VERSION : 0.1
   VAR_INPUT
      Zone : Int;
      ZonePos : Int;
      ClearOfStopDist : Int;
   END_VAR
   VAR_OUTPUT
      CarrierNumber : Int;
      MoveFwdCommand : Bool;
      DriveCmdSpeed : Int;
      NextCarrierNum : Word;
      NextStopPosition : DWord;
      AtCmdPosition : Bool;
      CarrierInTransitToNextZone : Bool;
   END_VAR
   VAR
      PreviousCarrierNumMemory : Word;
      TrafficCopCarrierZnBuffer : Array[0..40] of "UDT_TrafficCop";
      LastCarrierNextZnPos : Int;
      CarNumZnPos : Int;
      NextZone : Int;
      EndPos_LowLimit : DWord;
      EndPos_HighLimit : DWord;
      ClrOfStopPos_LowLimit : DWord;
      ClrOfStopPos_HighLimit : DWord;
      ClearOfStopPos : DWord;
      ClearToMoveTrain : Bool;
      PrevZone : Int;
      PrevZone_CarrierReady : Bool;
      LastCarrierCurrentZnPos : Int;
      LastCarrierNumber : Word;
      CarrierInTransitToProdZone : Bool;
      ResetCarrierInTransToProd : Bool;
      WaitPositionMemory : DInt;
      OneShot : Bool;
      NextCarrierOffset : DWord;
      PrevZone_EndPos_LowLimit : DWord;
      PrevZone_EndPos_HighLimit : DWord;
   END_VAR
   VAR_TEMP
      NextZoneBuffer : Int;
      LastZone : Int;
      HighSpeedSetpoint : Word;
      LowSpeedSetpoint : Word;
      NextZonePosition : Int;
      NextCarrierOffsetSetup1 : UDInt;
      NextCarrierOffsetSetup2 : UDInt;
   END_VAR
   VAR_TEMP   // added for the SCL form of the ladder/FBD networks
      _w1 : Bool;
      _w2 : Bool;
      _w3 : Bool;
      _w4 : Bool;
      _w5 : Bool;
   END_VAR
BEGIN

REGION Network 1
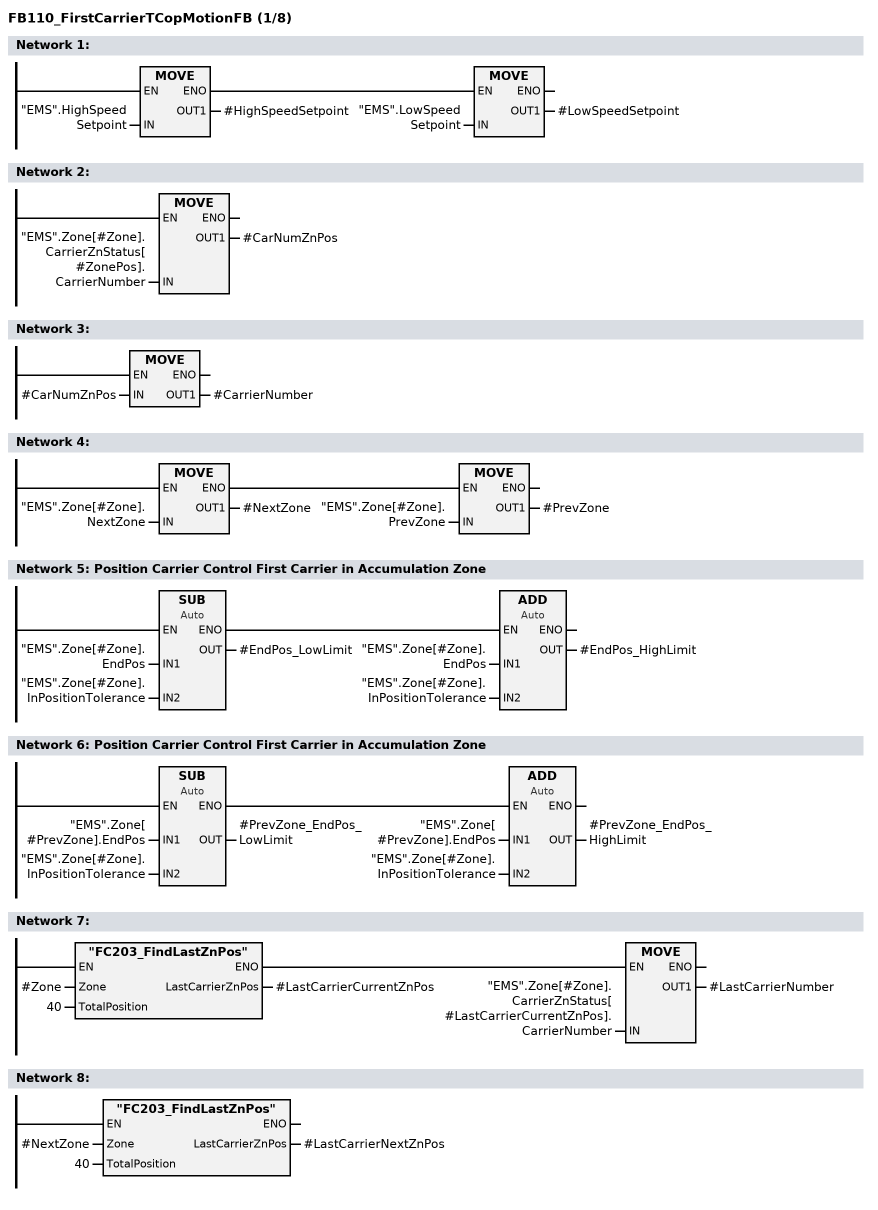
   RUNG wire#powerrail
      Move(in := "EMS".HighSpeedSetpoint, out1 => #HighSpeedSetpoint)
      Move(in := "EMS".LowSpeedSetpoint, out1 => #LowSpeedSetpoint)
   END_RUNG
   // the same network as SCL:
   #HighSpeedSetpoint := "EMS".HighSpeedSetpoint;
   #LowSpeedSetpoint := "EMS".LowSpeedSetpoint;
END_REGION

REGION Network 2
   RUNG wire#powerrail
      Move(in := "EMS".Zone[#Zone].CarrierZnStatus[#ZonePos].CarrierNumber, out1 => #CarNumZnPos)
   END_RUNG
   // the same network as SCL:
   #CarNumZnPos := "EMS".Zone[#Zone].CarrierZnStatus[#ZonePos].CarrierNumber;
END_REGION

REGION Network 3
   RUNG wire#powerrail
      Move(in := #CarNumZnPos, out1 => #CarrierNumber)
   END_RUNG
   // the same network as SCL:
   #CarrierNumber := #CarNumZnPos;
END_REGION

REGION Network 4
   RUNG wire#powerrail
      Move(in := "EMS".Zone[#Zone].NextZone, out1 => #NextZone)
      Move(in := "EMS".Zone[#Zone].PrevZone, out1 => #PrevZone)
   END_RUNG
   // the same network as SCL:
   #NextZone := "EMS".Zone[#Zone].NextZone;
   #PrevZone := "EMS".Zone[#Zone].PrevZone;
END_REGION

REGION Network 5: Position Carrier Control First Carrier in Accumulation Zone
   RUNG wire#powerrail
      Sub(in1 := "EMS".Zone[#Zone].EndPos, in2 := "EMS".Zone[#Zone].InPositionTolerance, out => #EndPos_LowLimit)
      Add(in1 := "EMS".Zone[#Zone].EndPos, in2 := "EMS".Zone[#Zone].InPositionTolerance, out => #EndPos_HighLimit)
   END_RUNG
   // the same network as SCL:
   #EndPos_LowLimit := "EMS".Zone[#Zone].EndPos - "EMS".Zone[#Zone].InPositionTolerance;
   #EndPos_HighLimit := "EMS".Zone[#Zone].EndPos + "EMS".Zone[#Zone].InPositionTolerance;
END_REGION

REGION Network 6: Position Carrier Control First Carrier in Accumulation Zone
   RUNG wire#powerrail
      Sub(in1 := "EMS".Zone[#PrevZone].EndPos, in2 := "EMS".Zone[#Zone].InPositionTolerance, out => #PrevZone_EndPos_LowLimit)
      Add(in1 := "EMS".Zone[#PrevZone].EndPos, in2 := "EMS".Zone[#Zone].InPositionTolerance, out => #PrevZone_EndPos_HighLimit)
   END_RUNG
   // the same network as SCL:
   #PrevZone_EndPos_LowLimit := "EMS".Zone[#PrevZone].EndPos - "EMS".Zone[#Zone].InPositionTolerance;
   #PrevZone_EndPos_HighLimit := "EMS".Zone[#PrevZone].EndPos + "EMS".Zone[#Zone].InPositionTolerance;
END_REGION

REGION Network 7
   RUNG wire#powerrail
      "FC203_FindLastZnPos"(Zone := #Zone, TotalPosition := 40, LastCarrierZnPos => #LastCarrierCurrentZnPos)
      Move(in := "EMS".Zone[#Zone].CarrierZnStatus[#LastCarrierCurrentZnPos].CarrierNumber, out1 => #LastCarrierNumber)
   END_RUNG
   // the same network as SCL:
   "FC203_FindLastZnPos"(Zone := #Zone,
                         TotalPosition := 40,
                         LastCarrierZnPos => #LastCarrierCurrentZnPos,
                         ENO => #_w1);
   IF #_w1 THEN
       #LastCarrierNumber := "EMS".Zone[#Zone].CarrierZnStatus[#LastCarrierCurrentZnPos].CarrierNumber;
   END_IF;
END_REGION

REGION Network 8
   RUNG wire#powerrail
      "FC203_FindLastZnPos"(Zone := #NextZone, TotalPosition := 40, LastCarrierZnPos => #LastCarrierNextZnPos)
   END_RUNG
   // the same network as SCL:
   "FC203_FindLastZnPos"(Zone := #NextZone, TotalPosition := 40, LastCarrierZnPos => #LastCarrierNextZnPos);
END_REGION

REGION Network 9: Position Carrier Control First Carrier in Production Zone
   // Control of First Carrier in Zone Closest to end position/Stop.  Move command is issued to carrier. Carrier will move in auto.
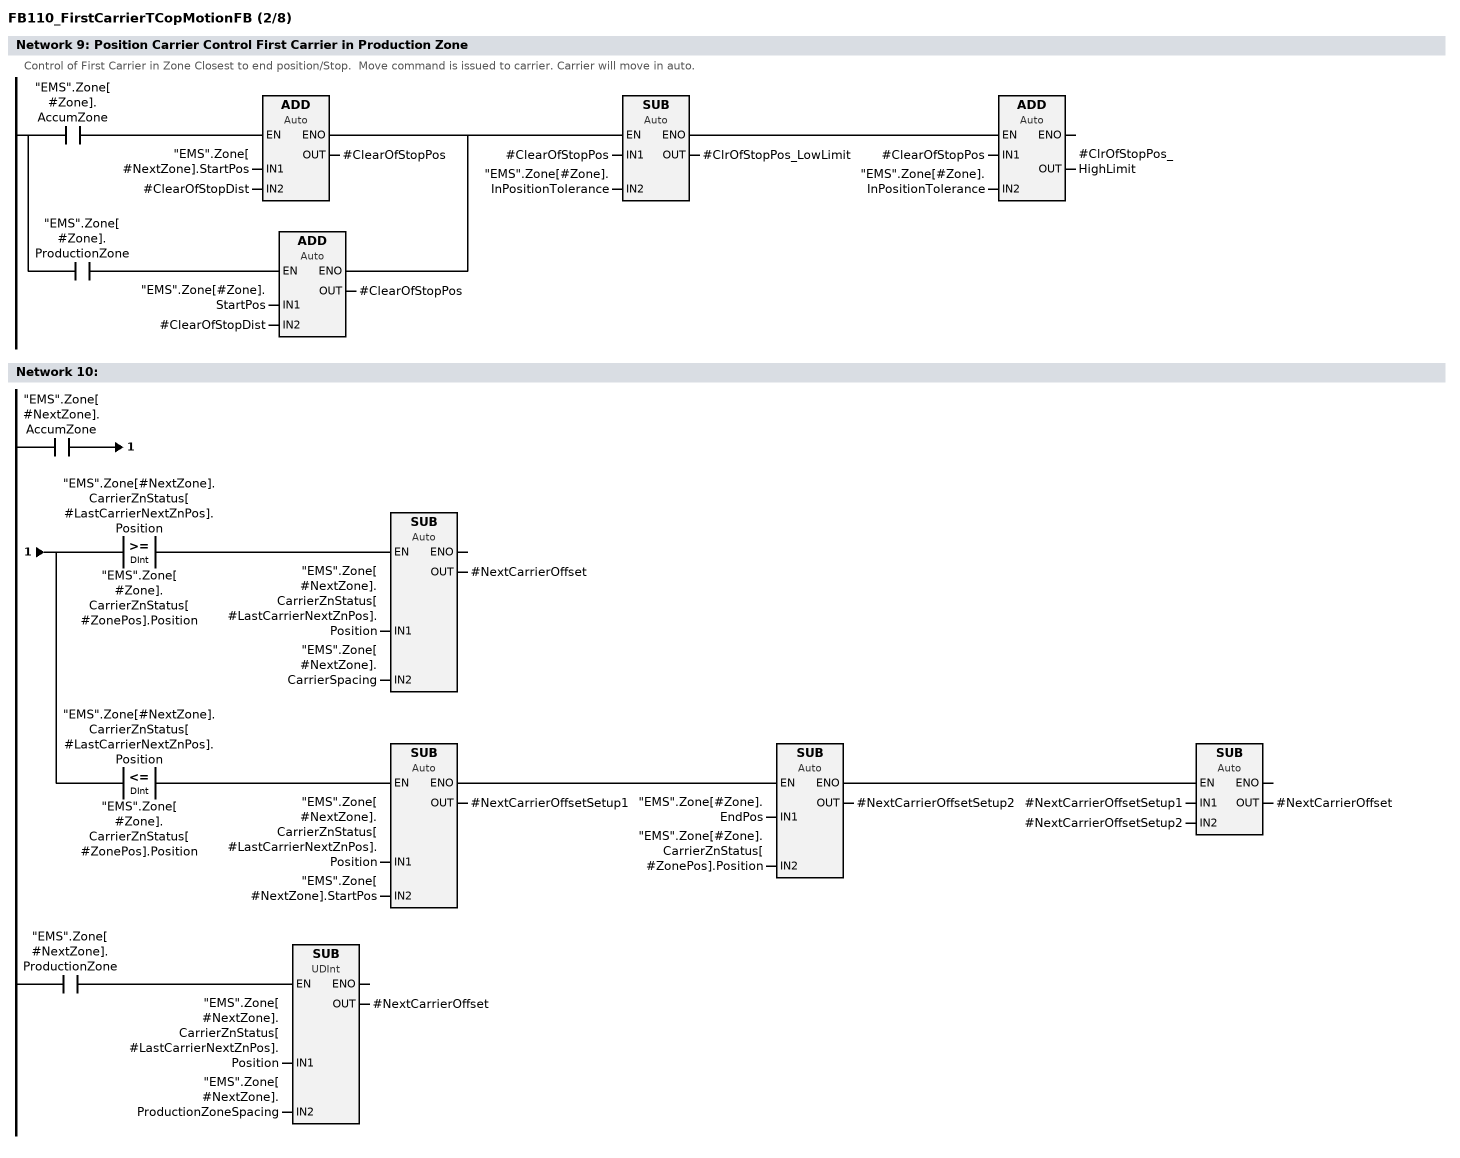
   RUNG wire#powerrail
      Contact( "EMS".Zone[#Zone].AccumZone )
      Add(in1 := "EMS".Zone[#NextZone].StartPos, in2 := #ClearOfStopDist, out => #ClearOfStopPos)
      wire#w1
      Sub(in1 := #ClearOfStopPos, in2 := "EMS".Zone[#Zone].InPositionTolerance, out => #ClrOfStopPos_LowLimit)
      Add(in1 := #ClearOfStopPos, in2 := "EMS".Zone[#Zone].InPositionTolerance, out => #ClrOfStopPos_HighLimit)
   END_RUNG
   RUNG wire#powerrail
      Contact( "EMS".Zone[#Zone].ProductionZone )
      Add(in1 := "EMS".Zone[#Zone].StartPos, in2 := #ClearOfStopDist, out => #ClearOfStopPos)
   END_RUNG wire#w1
   // the same network as SCL:
   IF "EMS".Zone[#Zone].AccumZone THEN
       #ClearOfStopPos := "EMS".Zone[#NextZone].StartPos + #ClearOfStopDist;
   END_IF;
   IF "EMS".Zone[#Zone].ProductionZone THEN
       #ClearOfStopPos := "EMS".Zone[#Zone].StartPos + #ClearOfStopDist;
   END_IF;
   IF "EMS".Zone[#Zone].AccumZone OR "EMS".Zone[#Zone].ProductionZone THEN
       #ClrOfStopPos_LowLimit := #ClearOfStopPos - "EMS".Zone[#Zone].InPositionTolerance;
       #ClrOfStopPos_HighLimit := #ClearOfStopPos + "EMS".Zone[#Zone].InPositionTolerance;
   END_IF;
END_REGION

REGION Network 10
   RUNG wire#powerrail
      Contact( "EMS".Zone[#NextZone].AccumZone )
      wire#w1
      { S7_Templates := "SrcType := DInt" } GE_Contact(in1 := "EMS".Zone[#NextZone].CarrierZnStatus[#LastCarrierNextZnPos].Position, in2 := "EMS".Zone[#Zone].CarrierZnStatus[#ZonePos].Position)
      Sub(in1 := "EMS".Zone[#NextZone].CarrierZnStatus[#LastCarrierNextZnPos].Position, in2 := "EMS".Zone[#NextZone].CarrierSpacing, out => #NextCarrierOffset)
   END_RUNG
   RUNG wire#w1
      { S7_Templates := "SrcType := DInt" } LE_Contact(in1 := "EMS".Zone[#NextZone].CarrierZnStatus[#LastCarrierNextZnPos].Position, in2 := "EMS".Zone[#Zone].CarrierZnStatus[#ZonePos].Position)
      Sub(in1 := "EMS".Zone[#NextZone].CarrierZnStatus[#LastCarrierNextZnPos].Position, in2 := "EMS".Zone[#NextZone].StartPos, out => #NextCarrierOffsetSetup1)
      Sub(in1 := "EMS".Zone[#Zone].EndPos, in2 := "EMS".Zone[#Zone].CarrierZnStatus[#ZonePos].Position, out => #NextCarrierOffsetSetup2)
      Sub(in1 := #NextCarrierOffsetSetup1, in2 := #NextCarrierOffsetSetup2, out => #NextCarrierOffset)
   END_RUNG
   RUNG wire#powerrail
      Contact( "EMS".Zone[#NextZone].ProductionZone )
      { S7_Templates := "SrcType := UDInt" } Sub(in1 := "EMS".Zone[#NextZone].CarrierZnStatus[#LastCarrierNextZnPos].Position, in2 := "EMS".Zone[#NextZone].ProductionZoneSpacing, out => #NextCarrierOffset)
   END_RUNG
   // the same network as SCL:
   IF "EMS".Zone[#NextZone].AccumZone AND ("EMS".Zone[#NextZone].CarrierZnStatus[#LastCarrierNextZnPos].Position >= "EMS".Zone[#Zone].CarrierZnStatus[#ZonePos].Position) THEN
       #NextCarrierOffset := "EMS".Zone[#NextZone].CarrierZnStatus[#LastCarrierNextZnPos].Position - "EMS".Zone[#NextZone].CarrierSpacing;
   END_IF;
   IF "EMS".Zone[#NextZone].AccumZone AND ("EMS".Zone[#NextZone].CarrierZnStatus[#LastCarrierNextZnPos].Position <= "EMS".Zone[#Zone].CarrierZnStatus[#ZonePos].Position) THEN
       #NextCarrierOffsetSetup1 := "EMS".Zone[#NextZone].CarrierZnStatus[#LastCarrierNextZnPos].Position - "EMS".Zone[#NextZone].StartPos;
       #NextCarrierOffsetSetup2 := "EMS".Zone[#Zone].EndPos - "EMS".Zone[#Zone].CarrierZnStatus[#ZonePos].Position;
       #NextCarrierOffset := #NextCarrierOffsetSetup1 - #NextCarrierOffsetSetup2;
   END_IF;
   IF "EMS".Zone[#NextZone].ProductionZone THEN
       #NextCarrierOffset := "EMS".Zone[#NextZone].CarrierZnStatus[#LastCarrierNextZnPos].Position - "EMS".Zone[#NextZone].ProductionZoneSpacing;
   END_IF;
END_REGION

REGION Network 11
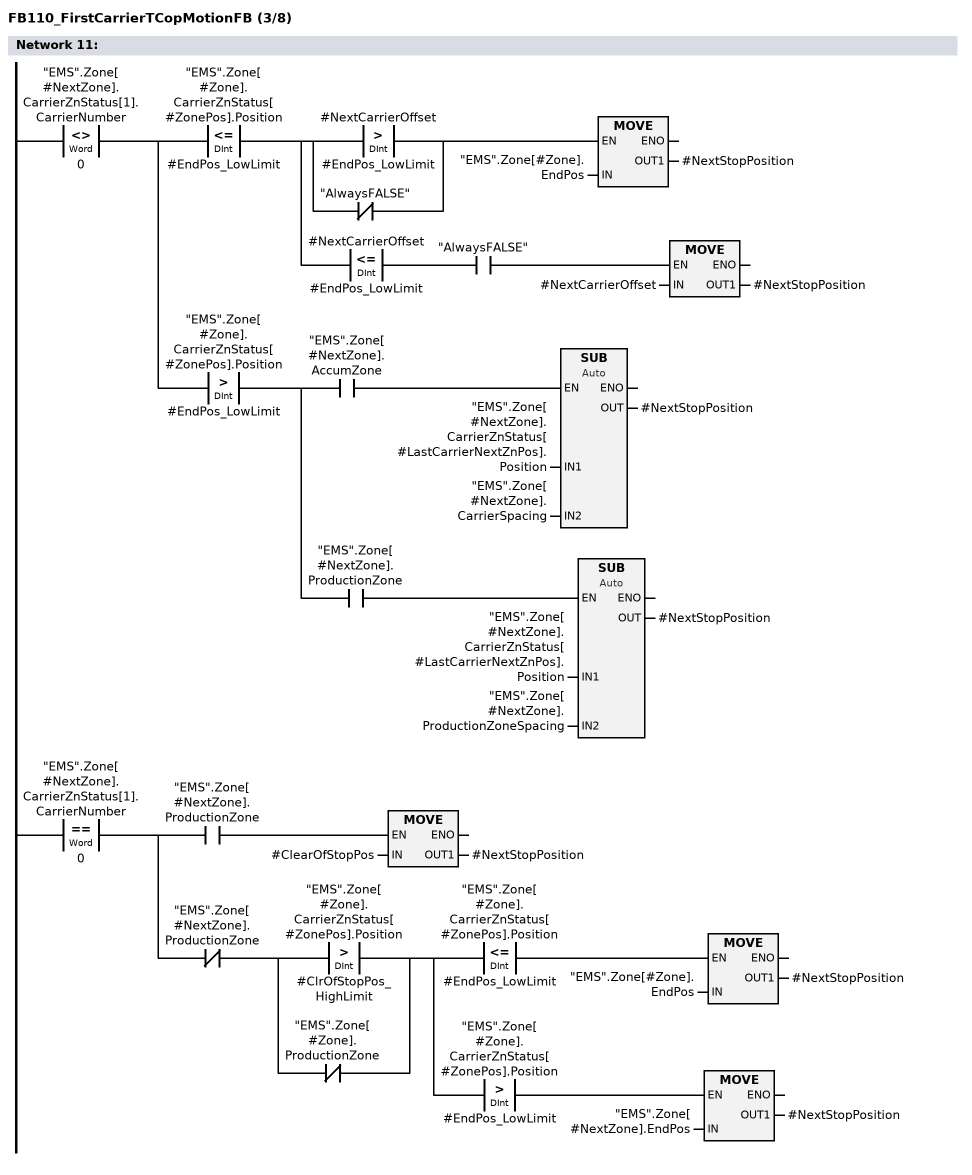
   RUNG wire#powerrail
      { S7_Templates := "SrcType := Word" } NE_Contact(in1 := "EMS".Zone[#NextZone].CarrierZnStatus[1].CarrierNumber, in2 := 0)
      wire#w1
      { S7_Templates := "SrcType := DInt" } LE_Contact(in1 := "EMS".Zone[#Zone].CarrierZnStatus[#ZonePos].Position, in2 := #EndPos_LowLimit)
      wire#w2
      { S7_Templates := "SrcType := DInt" } GT_Contact(in1 := #NextCarrierOffset, in2 := #EndPos_LowLimit)
      wire#w3
      Move(in := "EMS".Zone[#Zone].EndPos, out1 => #NextStopPosition)
   END_RUNG
   RUNG wire#w2
      I_Contact( "AlwaysFALSE" )
   END_RUNG wire#w3
   RUNG wire#w2
      { S7_Templates := "SrcType := DInt" } LE_Contact(in1 := #NextCarrierOffset, in2 := #EndPos_LowLimit)
      Contact( "AlwaysFALSE" )
      Move(in := #NextCarrierOffset, out1 => #NextStopPosition)
   END_RUNG
   RUNG wire#w1
      { S7_Templates := "SrcType := DInt" } GT_Contact(in1 := "EMS".Zone[#Zone].CarrierZnStatus[#ZonePos].Position, in2 := #EndPos_LowLimit)
      wire#w4
      Contact( "EMS".Zone[#NextZone].AccumZone )
      Sub(in1 := "EMS".Zone[#NextZone].CarrierZnStatus[#LastCarrierNextZnPos].Position, in2 := "EMS".Zone[#NextZone].CarrierSpacing, out => #NextStopPosition)
   END_RUNG
   RUNG wire#w4
      Contact( "EMS".Zone[#NextZone].ProductionZone )
      Sub(in1 := "EMS".Zone[#NextZone].CarrierZnStatus[#LastCarrierNextZnPos].Position, in2 := "EMS".Zone[#NextZone].ProductionZoneSpacing, out => #NextStopPosition)
   END_RUNG
   RUNG wire#powerrail
      { S7_Templates := "SrcType := Word" } EQ_Contact(in1 := "EMS".Zone[#NextZone].CarrierZnStatus[1].CarrierNumber, in2 := 0)
      wire#w5
      Contact( "EMS".Zone[#NextZone].ProductionZone )
      Move(in := #ClearOfStopPos, out1 => #NextStopPosition)
   END_RUNG
   RUNG wire#w5
      I_Contact( "EMS".Zone[#NextZone].ProductionZone )
      wire#w6
      { S7_Templates := "SrcType := DInt" } GT_Contact(in1 := "EMS".Zone[#Zone].CarrierZnStatus[#ZonePos].Position, in2 := #ClrOfStopPos_HighLimit)
      wire#w7
      { S7_Templates := "SrcType := DInt" } LE_Contact(in1 := "EMS".Zone[#Zone].CarrierZnStatus[#ZonePos].Position, in2 := #EndPos_LowLimit)
      Move(in := "EMS".Zone[#Zone].EndPos, out1 => #NextStopPosition)
   END_RUNG
   RUNG wire#w6
      I_Contact( "EMS".Zone[#Zone].ProductionZone )
   END_RUNG wire#w7
   RUNG wire#w7
      { S7_Templates := "SrcType := DInt" } GT_Contact(in1 := "EMS".Zone[#Zone].CarrierZnStatus[#ZonePos].Position, in2 := #EndPos_LowLimit)
      Move(in := "EMS".Zone[#NextZone].EndPos, out1 => #NextStopPosition)
   END_RUNG
   // the same network as SCL:
   #_w1 := "EMS".Zone[#NextZone].CarrierZnStatus[1].CarrierNumber <> 0;
   #_w2 := #_w1 AND ("EMS".Zone[#Zone].CarrierZnStatus[#ZonePos].Position <= #EndPos_LowLimit);
   IF #_w2 AND ((#NextCarrierOffset > #EndPos_LowLimit) OR NOT "AlwaysFALSE") THEN
       #NextStopPosition := "EMS".Zone[#Zone].EndPos;
   END_IF;
   IF #_w2 AND (#NextCarrierOffset <= #EndPos_LowLimit) AND "AlwaysFALSE" THEN
       #NextStopPosition := #NextCarrierOffset;
   END_IF;
   #_w3 := #_w1 AND ("EMS".Zone[#Zone].CarrierZnStatus[#ZonePos].Position > #EndPos_LowLimit);
   IF #_w3 AND "EMS".Zone[#NextZone].AccumZone THEN
       #NextStopPosition := "EMS".Zone[#NextZone].CarrierZnStatus[#LastCarrierNextZnPos].Position - "EMS".Zone[#NextZone].CarrierSpacing;
   END_IF;
   IF #_w3 AND "EMS".Zone[#NextZone].ProductionZone THEN
       #NextStopPosition := "EMS".Zone[#NextZone].CarrierZnStatus[#LastCarrierNextZnPos].Position - "EMS".Zone[#NextZone].ProductionZoneSpacing;
   END_IF;
   #_w4 := "EMS".Zone[#NextZone].CarrierZnStatus[1].CarrierNumber = 0;
   IF #_w4 AND "EMS".Zone[#NextZone].ProductionZone THEN #NextStopPosition := #ClearOfStopPos; END_IF;
   #_w5 := #_w4 AND NOT "EMS".Zone[#NextZone].ProductionZone AND (("EMS".Zone[#Zone].CarrierZnStatus[#ZonePos].Position > #ClrOfStopPos_HighLimit) OR NOT "EMS".Zone[#Zone].ProductionZone);
   IF #_w5 AND ("EMS".Zone[#Zone].CarrierZnStatus[#ZonePos].Position <= #EndPos_LowLimit) THEN
       #NextStopPosition := "EMS".Zone[#Zone].EndPos;
   END_IF;
   IF #_w5 AND ("EMS".Zone[#Zone].CarrierZnStatus[#ZonePos].Position > #EndPos_LowLimit) THEN
       #NextStopPosition := "EMS".Zone[#NextZone].EndPos;
   END_IF;
END_REGION

REGION Network 12
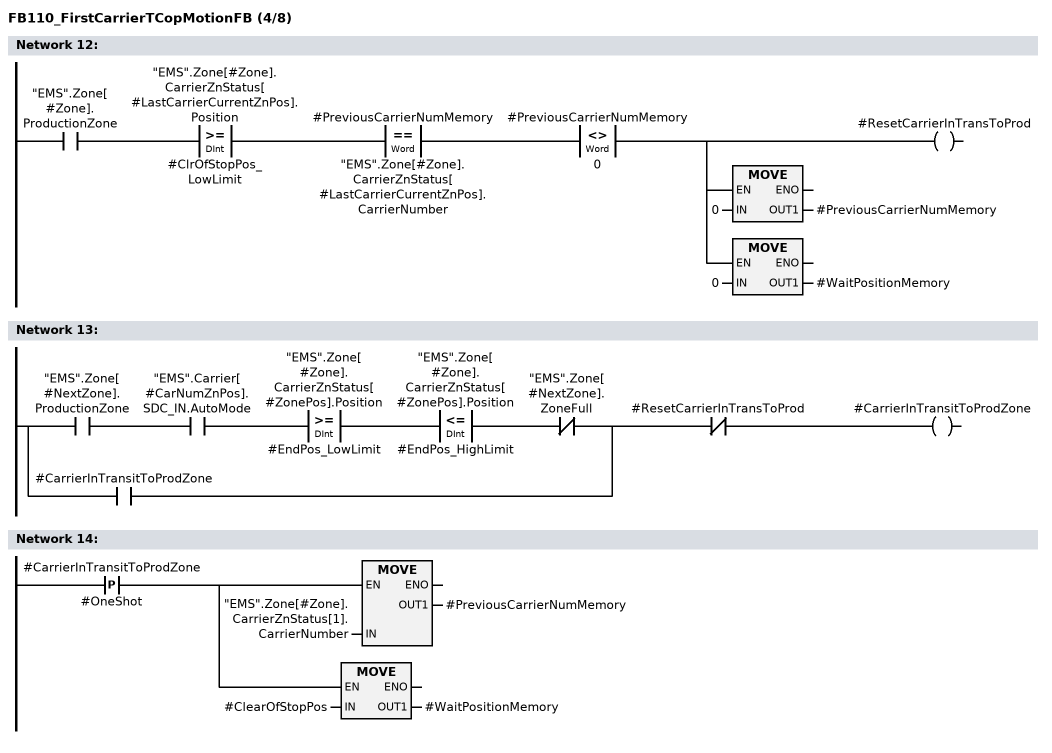
   RUNG wire#powerrail
      Contact( "EMS".Zone[#Zone].ProductionZone )
      { S7_Templates := "SrcType := DInt" } GE_Contact(in1 := "EMS".Zone[#Zone].CarrierZnStatus[#LastCarrierCurrentZnPos].Position, in2 := #ClrOfStopPos_LowLimit)
      { S7_Templates := "SrcType := Word" } EQ_Contact(in1 := #PreviousCarrierNumMemory, in2 := "EMS".Zone[#Zone].CarrierZnStatus[#LastCarrierCurrentZnPos].CarrierNumber)
      { S7_Templates := "SrcType := Word" } NE_Contact(in1 := #PreviousCarrierNumMemory, in2 := 0)
      wire#w1
      Coil( #ResetCarrierInTransToProd )
   END_RUNG
   RUNG wire#w1
      Move(in := 0, out1 => #PreviousCarrierNumMemory)
   END_RUNG
   RUNG wire#w1
      Move(in := 0, out1 => #WaitPositionMemory)
   END_RUNG
   // the same network as SCL:
   #ResetCarrierInTransToProd := "EMS".Zone[#Zone].ProductionZone AND ("EMS".Zone[#Zone].CarrierZnStatus[#LastCarrierCurrentZnPos].Position >= #ClrOfStopPos_LowLimit) AND (#PreviousCarrierNumMemory = "EMS".Zone[#Zone].CarrierZnStatus[#LastCarrierCurrentZnPos].CarrierNumber) AND (#PreviousCarrierNumMemory <> 0);
   IF #ResetCarrierInTransToProd THEN
       #PreviousCarrierNumMemory := 0;
       #WaitPositionMemory := 0;
   END_IF;
END_REGION

REGION Network 13
   RUNG wire#powerrail
      Contact( "EMS".Zone[#NextZone].ProductionZone )
      Contact( "EMS".Carrier[#CarNumZnPos].SDC_IN.AutoMode )
      { S7_Templates := "SrcType := DInt" } GE_Contact(in1 := "EMS".Zone[#Zone].CarrierZnStatus[#ZonePos].Position, in2 := #EndPos_LowLimit)
      { S7_Templates := "SrcType := DInt" } LE_Contact(in1 := "EMS".Zone[#Zone].CarrierZnStatus[#ZonePos].Position, in2 := #EndPos_HighLimit)
      I_Contact( "EMS".Zone[#NextZone].ZoneFull )
      wire#w1
      I_Contact( #ResetCarrierInTransToProd )
      Coil( #CarrierInTransitToProdZone )
   END_RUNG
   RUNG wire#powerrail
      Contact( #CarrierInTransitToProdZone )
   END_RUNG wire#w1
   // the same network as SCL:
   #CarrierInTransitToProdZone := (("EMS".Zone[#NextZone].ProductionZone AND "EMS".Carrier[#CarNumZnPos].SDC_IN.AutoMode AND ("EMS".Zone[#Zone].CarrierZnStatus[#ZonePos].Position >= #EndPos_LowLimit) AND ("EMS".Zone[#Zone].CarrierZnStatus[#ZonePos].Position <= #EndPos_HighLimit) AND NOT "EMS".Zone[#NextZone].ZoneFull) OR #CarrierInTransitToProdZone) AND NOT #ResetCarrierInTransToProd;
END_REGION

REGION Network 14
   RUNG wire#powerrail
      P_Contact(operand := #CarrierInTransitToProdZone, bit := #OneShot)
      wire#w1
      Move(in := "EMS".Zone[#Zone].CarrierZnStatus[1].CarrierNumber, out1 => #PreviousCarrierNumMemory)
   END_RUNG
   RUNG wire#w1
      Move(in := #ClearOfStopPos, out1 => #WaitPositionMemory)
   END_RUNG
   // the same network as SCL:
   #_w1 := #CarrierInTransitToProdZone AND NOT #OneShot;   // rising edge of #CarrierInTransitToProdZone
   #OneShot := #CarrierInTransitToProdZone;
   IF #_w1 THEN
       #PreviousCarrierNumMemory := "EMS".Zone[#Zone].CarrierZnStatus[1].CarrierNumber;
       #WaitPositionMemory := #ClearOfStopPos;
   END_IF;
END_REGION

REGION Network 15: Position Carrier Control First Carrier in Accumulation Zone
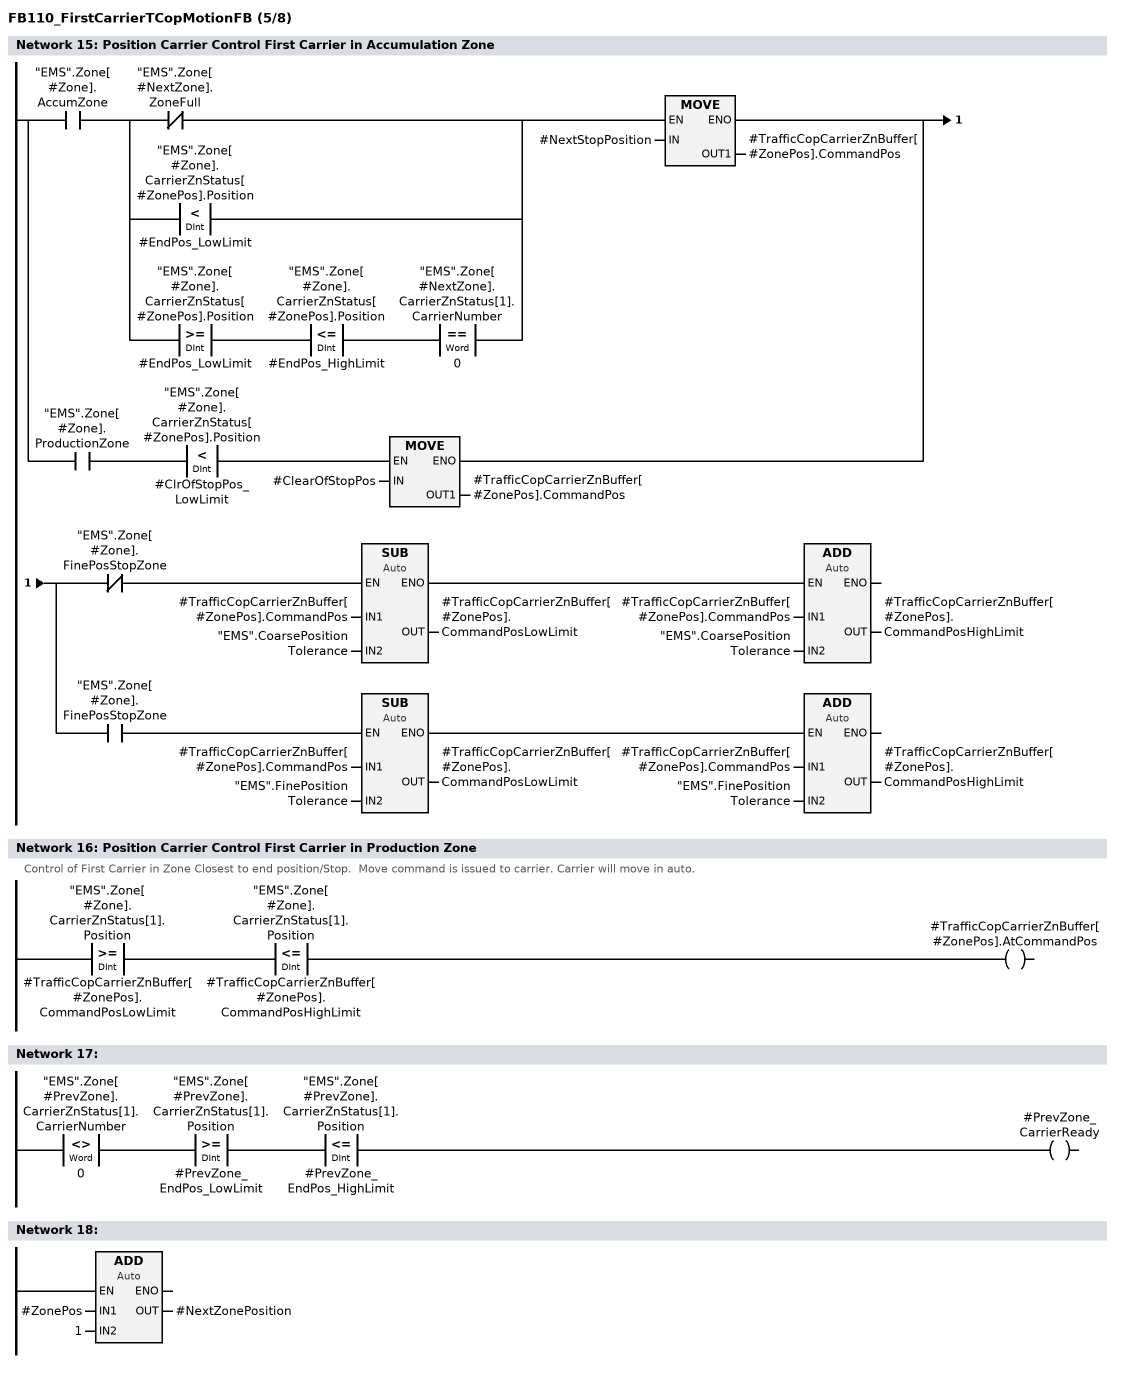
   RUNG wire#powerrail
      Contact( "EMS".Zone[#Zone].AccumZone )
      wire#w1
      I_Contact( "EMS".Zone[#NextZone].ZoneFull )
      wire#w2
      Move(in := #NextStopPosition, out1 => #TrafficCopCarrierZnBuffer[#ZonePos].CommandPos)
      wire#w3
      I_Contact( "EMS".Zone[#Zone].FinePosStopZone )
      Sub(in1 := #TrafficCopCarrierZnBuffer[#ZonePos].CommandPos, in2 := "EMS".CoarsePositionTolerance, out => #TrafficCopCarrierZnBuffer[#ZonePos].CommandPosLowLimit)
      Add(in1 := #TrafficCopCarrierZnBuffer[#ZonePos].CommandPos, in2 := "EMS".CoarsePositionTolerance, out => #TrafficCopCarrierZnBuffer[#ZonePos].CommandPosHighLimit)
   END_RUNG
   RUNG wire#w1
      { S7_Templates := "SrcType := DInt" } LT_Contact(in1 := "EMS".Zone[#Zone].CarrierZnStatus[#ZonePos].Position, in2 := #EndPos_LowLimit)
   END_RUNG wire#w2
   RUNG wire#w1
      { S7_Templates := "SrcType := DInt" } GE_Contact(in1 := "EMS".Zone[#Zone].CarrierZnStatus[#ZonePos].Position, in2 := #EndPos_LowLimit)
      { S7_Templates := "SrcType := DInt" } LE_Contact(in1 := "EMS".Zone[#Zone].CarrierZnStatus[#ZonePos].Position, in2 := #EndPos_HighLimit)
      { S7_Templates := "SrcType := Word" } EQ_Contact(in1 := "EMS".Zone[#NextZone].CarrierZnStatus[1].CarrierNumber, in2 := 0)
   END_RUNG wire#w2
   RUNG wire#powerrail
      Contact( "EMS".Zone[#Zone].ProductionZone )
      { S7_Templates := "SrcType := DInt" } LT_Contact(in1 := "EMS".Zone[#Zone].CarrierZnStatus[#ZonePos].Position, in2 := #ClrOfStopPos_LowLimit)
      Move(in := #ClearOfStopPos, out1 => #TrafficCopCarrierZnBuffer[#ZonePos].CommandPos)
   END_RUNG wire#w3
   RUNG wire#w3
      Contact( "EMS".Zone[#Zone].FinePosStopZone )
      Sub(in1 := #TrafficCopCarrierZnBuffer[#ZonePos].CommandPos, in2 := "EMS".FinePositionTolerance, out => #TrafficCopCarrierZnBuffer[#ZonePos].CommandPosLowLimit)
      Add(in1 := #TrafficCopCarrierZnBuffer[#ZonePos].CommandPos, in2 := "EMS".FinePositionTolerance, out => #TrafficCopCarrierZnBuffer[#ZonePos].CommandPosHighLimit)
   END_RUNG
   // the same network as SCL:
   #_w1 := "EMS".Zone[#Zone].AccumZone AND (NOT "EMS".Zone[#NextZone].ZoneFull OR ("EMS".Zone[#Zone].CarrierZnStatus[#ZonePos].Position < #EndPos_LowLimit) OR (("EMS".Zone[#Zone].CarrierZnStatus[#ZonePos].Position >= #EndPos_LowLimit) AND ("EMS".Zone[#Zone].CarrierZnStatus[#ZonePos].Position <= #EndPos_HighLimit) AND ("EMS".Zone[#NextZone].CarrierZnStatus[1].CarrierNumber = 0)));
   IF #_w1 THEN #TrafficCopCarrierZnBuffer[#ZonePos].CommandPos := #NextStopPosition; END_IF;
   #_w2 := "EMS".Zone[#Zone].ProductionZone AND ("EMS".Zone[#Zone].CarrierZnStatus[#ZonePos].Position < #ClrOfStopPos_LowLimit);
   IF #_w2 THEN #TrafficCopCarrierZnBuffer[#ZonePos].CommandPos := #ClearOfStopPos; END_IF;
   #_w3 := #_w1 OR #_w2;
   IF #_w3 AND NOT "EMS".Zone[#Zone].FinePosStopZone THEN
       #TrafficCopCarrierZnBuffer[#ZonePos].CommandPosLowLimit := #TrafficCopCarrierZnBuffer[#ZonePos].CommandPos - "EMS".CoarsePositionTolerance;
       #TrafficCopCarrierZnBuffer[#ZonePos].CommandPosHighLimit := #TrafficCopCarrierZnBuffer[#ZonePos].CommandPos + "EMS".CoarsePositionTolerance;
   END_IF;
   IF #_w3 AND "EMS".Zone[#Zone].FinePosStopZone THEN
       #TrafficCopCarrierZnBuffer[#ZonePos].CommandPosLowLimit := #TrafficCopCarrierZnBuffer[#ZonePos].CommandPos - "EMS".FinePositionTolerance;
       #TrafficCopCarrierZnBuffer[#ZonePos].CommandPosHighLimit := #TrafficCopCarrierZnBuffer[#ZonePos].CommandPos + "EMS".FinePositionTolerance;
   END_IF;
END_REGION
